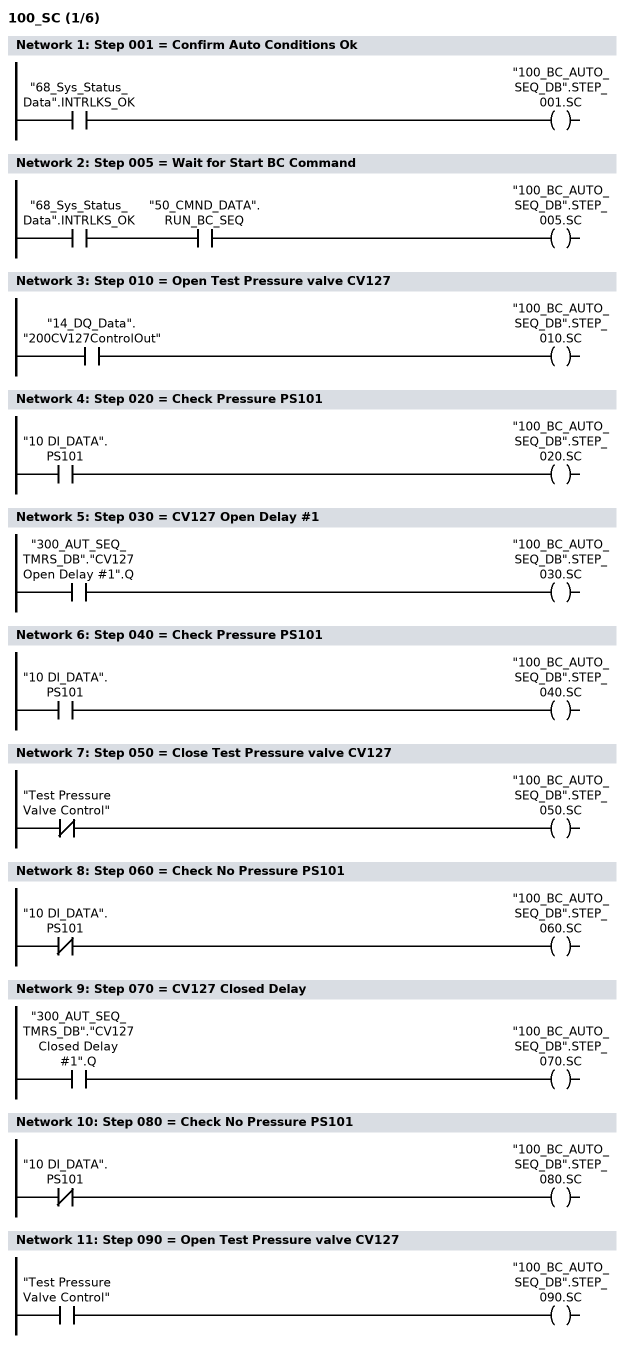
   RUNG wire#powerrail
      Contact( "68_Sys_Status_Data".INTRLKS_OK )
      Coil( "100_BC_AUTO_SEQ_DB".STEP_001.SC )
   END_RUNG
   // the same network as SCL:
   "100_BC_AUTO_SEQ_DB".STEP_001.SC := "68_Sys_Status_Data".INTRLKS_OK;
END_REGION

REGION Network 2: Step 005 = Wait for Start BC Command
   RUNG wire#powerrail
      Contact( "68_Sys_Status_Data".INTRLKS_OK )
      Contact( "50_CMND_DATA".RUN_BC_SEQ )
      Coil( "100_BC_AUTO_SEQ_DB".STEP_005.SC )
   END_RUNG
   // the same network as SCL:
   "100_BC_AUTO_SEQ_DB".STEP_005.SC := "68_Sys_Status_Data".INTRLKS_OK AND "50_CMND_DATA".RUN_BC_SEQ;
END_REGION

REGION Network 3: Step 010 = Open Test Pressure valve CV127
   RUNG wire#powerrail
      Contact( "14_DQ_Data"."200CV127ControlOut" )
      Coil( "100_BC_AUTO_SEQ_DB".STEP_010.SC )
   END_RUNG
   // the same network as SCL:
   "100_BC_AUTO_SEQ_DB".STEP_010.SC := "14_DQ_Data"."200CV127ControlOut";
END_REGION

REGION Network 4: Step 020 = Check Pressure PS101
   RUNG wire#powerrail
      Contact( "10 DI_DATA".PS101 )
      Coil( "100_BC_AUTO_SEQ_DB".STEP_020.SC )
   END_RUNG
   // the same network as SCL:
   "100_BC_AUTO_SEQ_DB".STEP_020.SC := "10 DI_DATA".PS101;
END_REGION

REGION Network 5: Step 030 = CV127 Open Delay #1
   RUNG wire#powerrail
      Contact( "300_AUT_SEQ_TMRS_DB"."CV127 Open Delay #1".Q )
      Coil( "100_BC_AUTO_SEQ_DB".STEP_030.SC )
   END_RUNG
   // the same network as SCL:
   "100_BC_AUTO_SEQ_DB".STEP_030.SC := "300_AUT_SEQ_TMRS_DB"."CV127 Open Delay #1".Q;
END_REGION

REGION Network 6: Step 040 = Check Pressure PS101
   RUNG wire#powerrail
      Contact( "10 DI_DATA".PS101 )
      Coil( "100_BC_AUTO_SEQ_DB".STEP_040.SC )
   END_RUNG
   // the same network as SCL:
   "100_BC_AUTO_SEQ_DB".STEP_040.SC := "10 DI_DATA".PS101;
END_REGION

REGION Network 7: Step 050 = Close Test Pressure valve CV127
   RUNG wire#powerrail
      I_Contact( "Test Pressure Valve Control" )
      Coil( "100_BC_AUTO_SEQ_DB".STEP_050.SC )
   END_RUNG
   // the same network as SCL:
   "100_BC_AUTO_SEQ_DB".STEP_050.SC := NOT "Test Pressure Valve Control";
END_REGION

REGION Network 8: Step 060 = Check No Pressure PS101
   RUNG wire#powerrail
      I_Contact( "10 DI_DATA".PS101 )
      Coil( "100_BC_AUTO_SEQ_DB".STEP_060.SC )
   END_RUNG
   // the same network as SCL:
   "100_BC_AUTO_SEQ_DB".STEP_060.SC := NOT "10 DI_DATA".PS101;
END_REGION

REGION Network 9: Step 070 = CV127 Closed Delay
   RUNG wire#powerrail
      Contact( "300_AUT_SEQ_TMRS_DB"."CV127 Closed Delay #1".Q )
      Coil( "100_BC_AUTO_SEQ_DB".STEP_070.SC )
   END_RUNG
   // the same network as SCL:
   "100_BC_AUTO_SEQ_DB".STEP_070.SC := "300_AUT_SEQ_TMRS_DB"."CV127 Closed Delay #1".Q;
END_REGION

REGION Network 10: Step 080 = Check No Pressure PS101
   RUNG wire#powerrail
      I_Contact( "10 DI_DATA".PS101 )
      Coil( "100_BC_AUTO_SEQ_DB".STEP_080.SC )
   END_RUNG
   // the same network as SCL:
   "100_BC_AUTO_SEQ_DB".STEP_080.SC := NOT "10 DI_DATA".PS101;
END_REGION

REGION Network 11: Step 090 = Open Test Pressure valve CV127
   RUNG wire#powerrail
      Contact( "Test Pressure Valve Control" )
      Coil( "100_BC_AUTO_SEQ_DB".STEP_090.SC )
   END_RUNG
   // the same network as SCL:
   "100_BC_AUTO_SEQ_DB".STEP_090.SC := "Test Pressure Valve Control";
END_REGION

REGION Network 12: Step 095 = Confirm CV403 Is Open
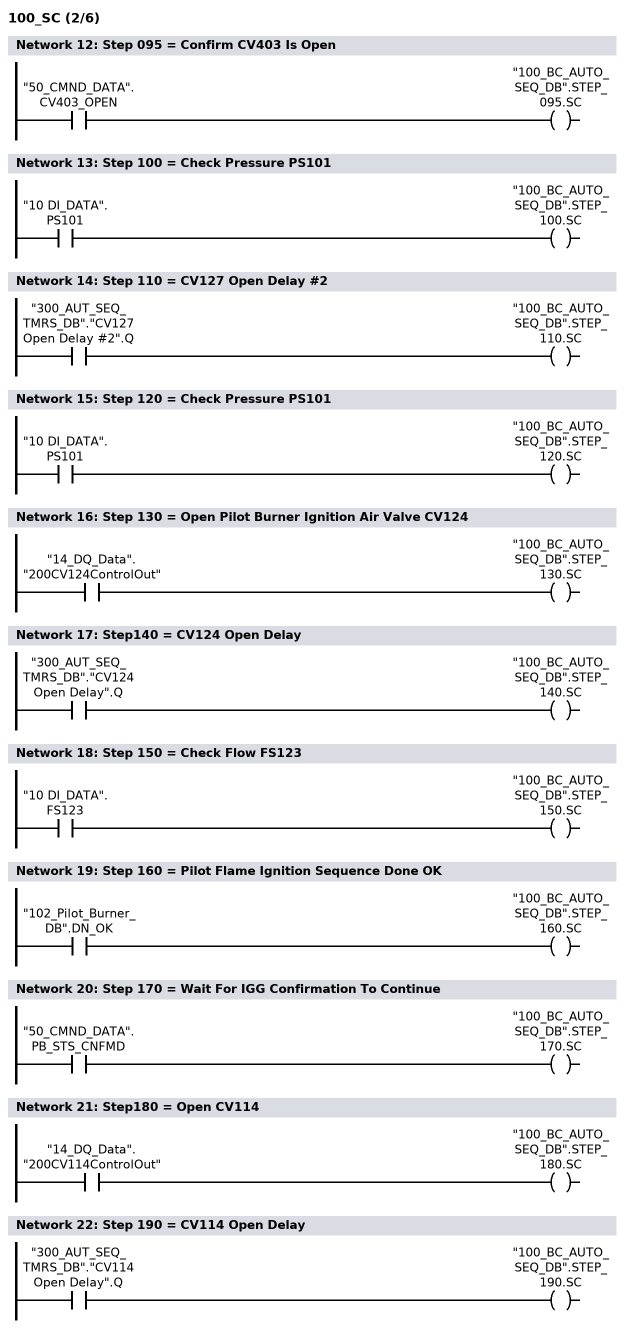
   RUNG wire#powerrail
      Contact( "50_CMND_DATA".CV403_OPEN )
      Coil( "100_BC_AUTO_SEQ_DB".STEP_095.SC )
   END_RUNG
   // the same network as SCL:
   "100_BC_AUTO_SEQ_DB".STEP_095.SC := "50_CMND_DATA".CV403_OPEN;
END_REGION

REGION Network 13: Step 100 = Check Pressure PS101
   RUNG wire#powerrail
      Contact( "10 DI_DATA".PS101 )
      Coil( "100_BC_AUTO_SEQ_DB".STEP_100.SC )
   END_RUNG
   // the same network as SCL:
   "100_BC_AUTO_SEQ_DB".STEP_100.SC := "10 DI_DATA".PS101;
END_REGION

REGION Network 14: Step 110 = CV127 Open Delay #2
   RUNG wire#powerrail
      Contact( "300_AUT_SEQ_TMRS_DB"."CV127 Open Delay #2".Q )
      Coil( "100_BC_AUTO_SEQ_DB".STEP_110.SC )
   END_RUNG
   // the same network as SCL:
   "100_BC_AUTO_SEQ_DB".STEP_110.SC := "300_AUT_SEQ_TMRS_DB"."CV127 Open Delay #2".Q;
END_REGION

REGION Network 15: Step 120 = Check Pressure PS101
   RUNG wire#powerrail
      Contact( "10 DI_DATA".PS101 )
      Coil( "100_BC_AUTO_SEQ_DB".STEP_120.SC )
   END_RUNG
   // the same network as SCL:
   "100_BC_AUTO_SEQ_DB".STEP_120.SC := "10 DI_DATA".PS101;
END_REGION

REGION Network 16: Step 130 = Open Pilot Burner Ignition Air Valve CV124
   RUNG wire#powerrail
      Contact( "14_DQ_Data"."200CV124ControlOut" )
      Coil( "100_BC_AUTO_SEQ_DB".STEP_130.SC )
   END_RUNG
   // the same network as SCL:
   "100_BC_AUTO_SEQ_DB".STEP_130.SC := "14_DQ_Data"."200CV124ControlOut";
END_REGION

REGION Network 17: Step140 = CV124 Open Delay
   RUNG wire#powerrail
      Contact( "300_AUT_SEQ_TMRS_DB"."CV124 Open Delay".Q )
      Coil( "100_BC_AUTO_SEQ_DB".STEP_140.SC )
   END_RUNG
   // the same network as SCL:
   "100_BC_AUTO_SEQ_DB".STEP_140.SC := "300_AUT_SEQ_TMRS_DB"."CV124 Open Delay".Q;
END_REGION

REGION Network 18: Step 150 = Check Flow FS123
   RUNG wire#powerrail
      Contact( "10 DI_DATA".FS123 )
      Coil( "100_BC_AUTO_SEQ_DB".STEP_150.SC )
   END_RUNG
   // the same network as SCL:
   "100_BC_AUTO_SEQ_DB".STEP_150.SC := "10 DI_DATA".FS123;
END_REGION

REGION Network 19: Step 160 = Pilot Flame Ignition Sequence Done OK
   RUNG wire#powerrail
      Contact( "102_Pilot_Burner_DB".DN_OK )
      Coil( "100_BC_AUTO_SEQ_DB".STEP_160.SC )
   END_RUNG
   // the same network as SCL:
   "100_BC_AUTO_SEQ_DB".STEP_160.SC := "102_Pilot_Burner_DB".DN_OK;
END_REGION

REGION Network 20: Step 170 = Wait For IGG Confirmation To Continue
   RUNG wire#powerrail
      Contact( "50_CMND_DATA".PB_STS_CNFMD )
      Coil( "100_BC_AUTO_SEQ_DB".STEP_170.SC )
   END_RUNG
   // the same network as SCL:
   "100_BC_AUTO_SEQ_DB".STEP_170.SC := "50_CMND_DATA".PB_STS_CNFMD;
END_REGION

REGION Network 21: Step180 = Open CV114
   RUNG wire#powerrail
      Contact( "14_DQ_Data"."200CV114ControlOut" )
      Coil( "100_BC_AUTO_SEQ_DB".STEP_180.SC )
   END_RUNG
   // the same network as SCL:
   "100_BC_AUTO_SEQ_DB".STEP_180.SC := "14_DQ_Data"."200CV114ControlOut";
END_REGION

REGION Network 22: Step 190 = CV114 Open Delay
   RUNG wire#powerrail
      Contact( "300_AUT_SEQ_TMRS_DB"."CV114 Open Delay".Q )
      Coil( "100_BC_AUTO_SEQ_DB".STEP_190.SC )
   END_RUNG
   // the same network as SCL:
   "100_BC_AUTO_SEQ_DB".STEP_190.SC := "300_AUT_SEQ_TMRS_DB"."CV114 Open Delay".Q;
END_REGION

REGION Network 23: Step 200 = Main Burner Ignition Sequence
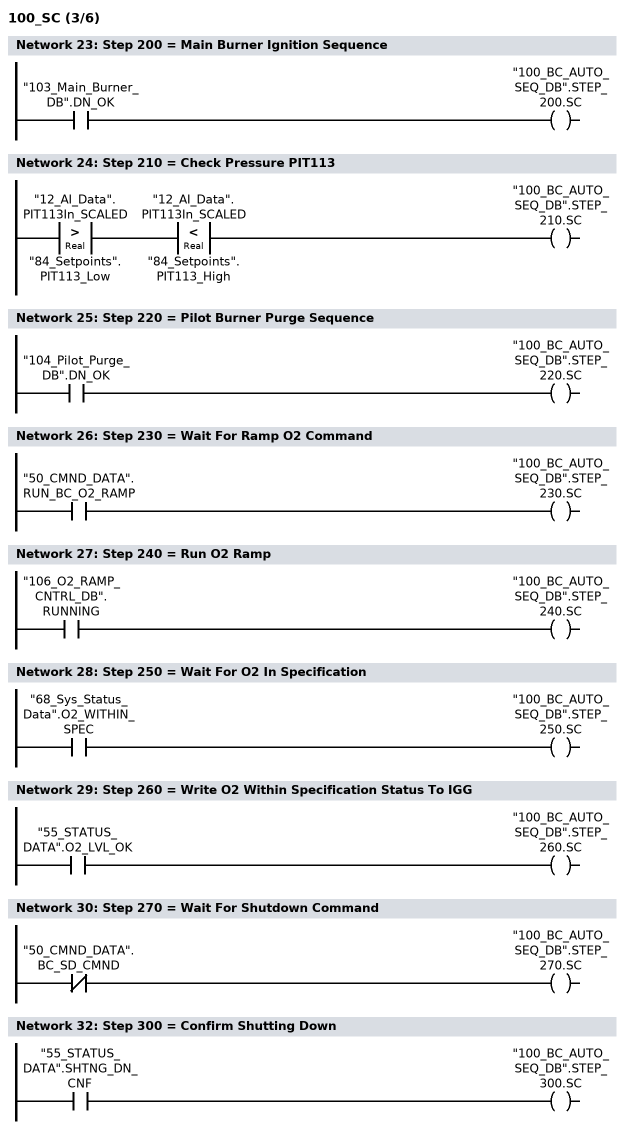
   RUNG wire#powerrail
      Contact( "103_Main_Burner_DB".DN_OK )
      Coil( "100_BC_AUTO_SEQ_DB".STEP_200.SC )
   END_RUNG
   // the same network as SCL:
   "100_BC_AUTO_SEQ_DB".STEP_200.SC := "103_Main_Burner_DB".DN_OK;
END_REGION

REGION Network 24: Step 210 = Check Pressure PIT113
   RUNG wire#powerrail
      { S7_Templates := "SrcType := Real" } GT_Contact(in1 := "12_AI_Data".PIT113In_SCALED, in2 := "84_Setpoints".PIT113_Low)
      { S7_Templates := "SrcType := Real" } LT_Contact(in1 := "12_AI_Data".PIT113In_SCALED, in2 := "84_Setpoints".PIT113_High)
      Coil( "100_BC_AUTO_SEQ_DB".STEP_210.SC )
   END_RUNG
   // the same network as SCL:
   "100_BC_AUTO_SEQ_DB".STEP_210.SC := ("12_AI_Data".PIT113In_SCALED > "84_Setpoints".PIT113_Low) AND ("12_AI_Data".PIT113In_SCALED < "84_Setpoints".PIT113_High);
END_REGION

REGION Network 25: Step 220 = Pilot Burner Purge Sequence
   RUNG wire#powerrail
      Contact( "104_Pilot_Purge_DB".DN_OK )
      Coil( "100_BC_AUTO_SEQ_DB".STEP_220.SC )
   END_RUNG
   // the same network as SCL:
   "100_BC_AUTO_SEQ_DB".STEP_220.SC := "104_Pilot_Purge_DB".DN_OK;
END_REGION

REGION Network 26: Step 230 = Wait For Ramp O2 Command
   RUNG wire#powerrail
      Contact( "50_CMND_DATA".RUN_BC_O2_RAMP )
      Coil( "100_BC_AUTO_SEQ_DB".STEP_230.SC )
   END_RUNG
   // the same network as SCL:
   "100_BC_AUTO_SEQ_DB".STEP_230.SC := "50_CMND_DATA".RUN_BC_O2_RAMP;
END_REGION

REGION Network 27: Step 240 = Run O2 Ramp
   RUNG wire#powerrail
      Contact( "106_O2_RAMP_CNTRL_DB".RUNNING )
      Coil( "100_BC_AUTO_SEQ_DB".STEP_240.SC )
   END_RUNG
   // the same network as SCL:
   "100_BC_AUTO_SEQ_DB".STEP_240.SC := "106_O2_RAMP_CNTRL_DB".RUNNING;
END_REGION

REGION Network 28: Step 250 = Wait For O2 In Specification
   RUNG wire#powerrail
      Contact( "68_Sys_Status_Data".O2_WITHIN_SPEC )
      Coil( "100_BC_AUTO_SEQ_DB".STEP_250.SC )
   END_RUNG
   // the same network as SCL:
   "100_BC_AUTO_SEQ_DB".STEP_250.SC := "68_Sys_Status_Data".O2_WITHIN_SPEC;
END_REGION

REGION Network 29: Step 260 = Write O2 Within Specification Status To IGG
   RUNG wire#powerrail
      Contact( "55_STATUS_DATA".O2_LVL_OK )
      Coil( "100_BC_AUTO_SEQ_DB".STEP_260.SC )
   END_RUNG
   // the same network as SCL:
   "100_BC_AUTO_SEQ_DB".STEP_260.SC := "55_STATUS_DATA".O2_LVL_OK;
END_REGION

REGION Network 30: Step 270 = Wait For Shutdown Command
   RUNG wire#powerrail
      I_Contact( "50_CMND_DATA".BC_SD_CMND )
      Coil( "100_BC_AUTO_SEQ_DB".STEP_270.SC )
   END_RUNG
   // the same network as SCL:
   "100_BC_AUTO_SEQ_DB".STEP_270.SC := NOT "50_CMND_DATA".BC_SD_CMND;
END_REGION

REGION Network 32: Step 300 = Confirm Shutting Down
   RUNG wire#powerrail
      Contact( "55_STATUS_DATA".SHTNG_DN_CNF )
      Coil( "100_BC_AUTO_SEQ_DB".STEP_300.SC )
   END_RUNG
   // the same network as SCL:
   "100_BC_AUTO_SEQ_DB".STEP_300.SC := "55_STATUS_DATA".SHTNG_DN_CNF;
END_REGION

REGION Network 33: Step 310 = CV203 To High O2 Standard Burn Setting
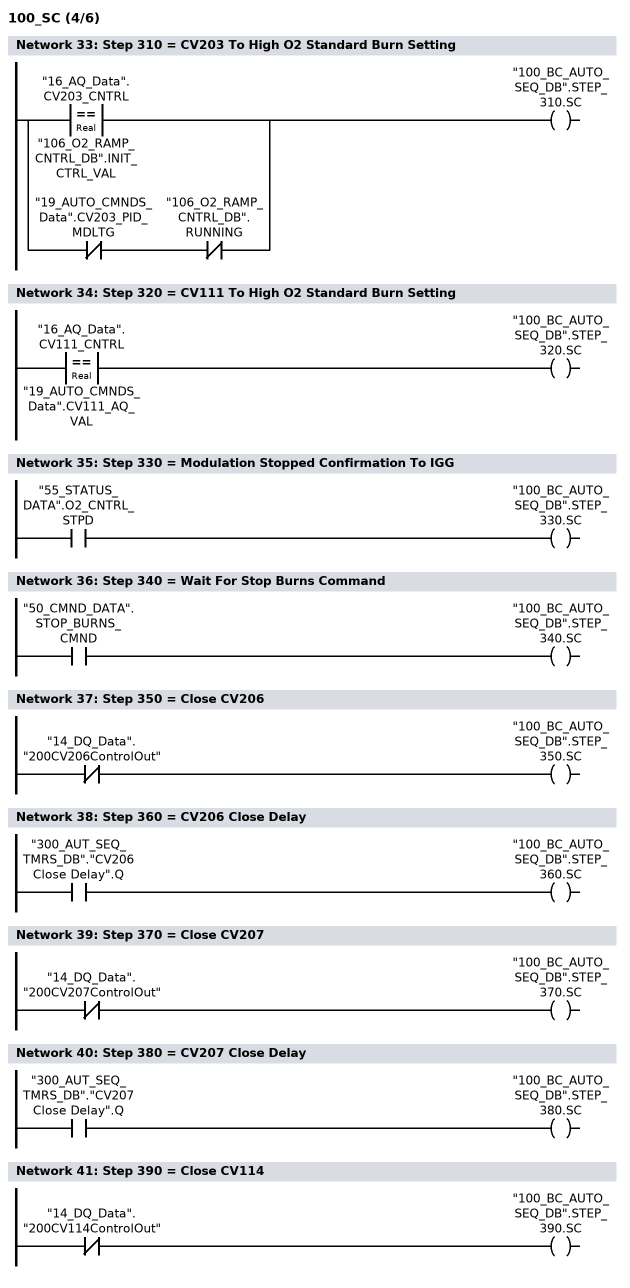
   RUNG wire#powerrail
      { S7_Templates := "SrcType := Real" } EQ_Contact(in1 := "16_AQ_Data".CV203_CNTRL, in2 := "106_O2_RAMP_CNTRL_DB".INIT_CTRL_VAL)
      wire#w1
      Coil( "100_BC_AUTO_SEQ_DB".STEP_310.SC )
   END_RUNG
   RUNG wire#powerrail
      I_Contact( "19_AUTO_CMNDS_Data".CV203_PID_MDLTG )
      I_Contact( "106_O2_RAMP_CNTRL_DB".RUNNING )
   END_RUNG wire#w1
   // the same network as SCL:
   "100_BC_AUTO_SEQ_DB".STEP_310.SC := ("16_AQ_Data".CV203_CNTRL = "106_O2_RAMP_CNTRL_DB".INIT_CTRL_VAL) OR (NOT "19_AUTO_CMNDS_Data".CV203_PID_MDLTG AND NOT "106_O2_RAMP_CNTRL_DB".RUNNING);
END_REGION

REGION Network 34: Step 320 = CV111 To High O2 Standard Burn Setting
   RUNG wire#powerrail
      { S7_Templates := "SrcType := Real" } EQ_Contact(in1 := "16_AQ_Data".CV111_CNTRL, in2 := "19_AUTO_CMNDS_Data".CV111_AQ_VAL)
      Coil( "100_BC_AUTO_SEQ_DB".STEP_320.SC )
   END_RUNG
   // the same network as SCL:
   "100_BC_AUTO_SEQ_DB".STEP_320.SC := "16_AQ_Data".CV111_CNTRL = "19_AUTO_CMNDS_Data".CV111_AQ_VAL;
END_REGION

REGION Network 35: Step 330 = Modulation Stopped Confirmation To IGG
   RUNG wire#powerrail
      Contact( "55_STATUS_DATA".O2_CNTRL_STPD )
      Coil( "100_BC_AUTO_SEQ_DB".STEP_330.SC )
   END_RUNG
   // the same network as SCL:
   "100_BC_AUTO_SEQ_DB".STEP_330.SC := "55_STATUS_DATA".O2_CNTRL_STPD;
END_REGION

REGION Network 36: Step 340 = Wait For Stop Burns Command
   RUNG wire#powerrail
      Contact( "50_CMND_DATA".STOP_BURNS_CMND )
      Coil( "100_BC_AUTO_SEQ_DB".STEP_340.SC )
   END_RUNG
   // the same network as SCL:
   "100_BC_AUTO_SEQ_DB".STEP_340.SC := "50_CMND_DATA".STOP_BURNS_CMND;
END_REGION

REGION Network 37: Step 350 = Close CV206
   RUNG wire#powerrail
      I_Contact( "14_DQ_Data"."200CV206ControlOut" )
      Coil( "100_BC_AUTO_SEQ_DB".STEP_350.SC )
   END_RUNG
   // the same network as SCL:
   "100_BC_AUTO_SEQ_DB".STEP_350.SC := NOT "14_DQ_Data"."200CV206ControlOut";
END_REGION

REGION Network 38: Step 360 = CV206 Close Delay
   RUNG wire#powerrail
      Contact( "300_AUT_SEQ_TMRS_DB"."CV206 Close Delay".Q )
      Coil( "100_BC_AUTO_SEQ_DB".STEP_360.SC )
   END_RUNG
   // the same network as SCL:
   "100_BC_AUTO_SEQ_DB".STEP_360.SC := "300_AUT_SEQ_TMRS_DB"."CV206 Close Delay".Q;
END_REGION

REGION Network 39: Step 370 = Close CV207
   RUNG wire#powerrail
      I_Contact( "14_DQ_Data"."200CV207ControlOut" )
      Coil( "100_BC_AUTO_SEQ_DB".STEP_370.SC )
   END_RUNG
   // the same network as SCL:
   "100_BC_AUTO_SEQ_DB".STEP_370.SC := NOT "14_DQ_Data"."200CV207ControlOut";
END_REGION

REGION Network 40: Step 380 = CV207 Close Delay
   RUNG wire#powerrail
      Contact( "300_AUT_SEQ_TMRS_DB"."CV207 Close Delay".Q )
      Coil( "100_BC_AUTO_SEQ_DB".STEP_380.SC )
   END_RUNG
   // the same network as SCL:
   "100_BC_AUTO_SEQ_DB".STEP_380.SC := "300_AUT_SEQ_TMRS_DB"."CV207 Close Delay".Q;
END_REGION

REGION Network 41: Step 390 = Close CV114
   RUNG wire#powerrail
      I_Contact( "14_DQ_Data"."200CV114ControlOut" )
      Coil( "100_BC_AUTO_SEQ_DB".STEP_390.SC )
   END_RUNG
   // the same network as SCL:
   "100_BC_AUTO_SEQ_DB".STEP_390.SC := NOT "14_DQ_Data"."200CV114ControlOut";
END_REGION

REGION Network 42: Step 400 = CV114 Close Delay
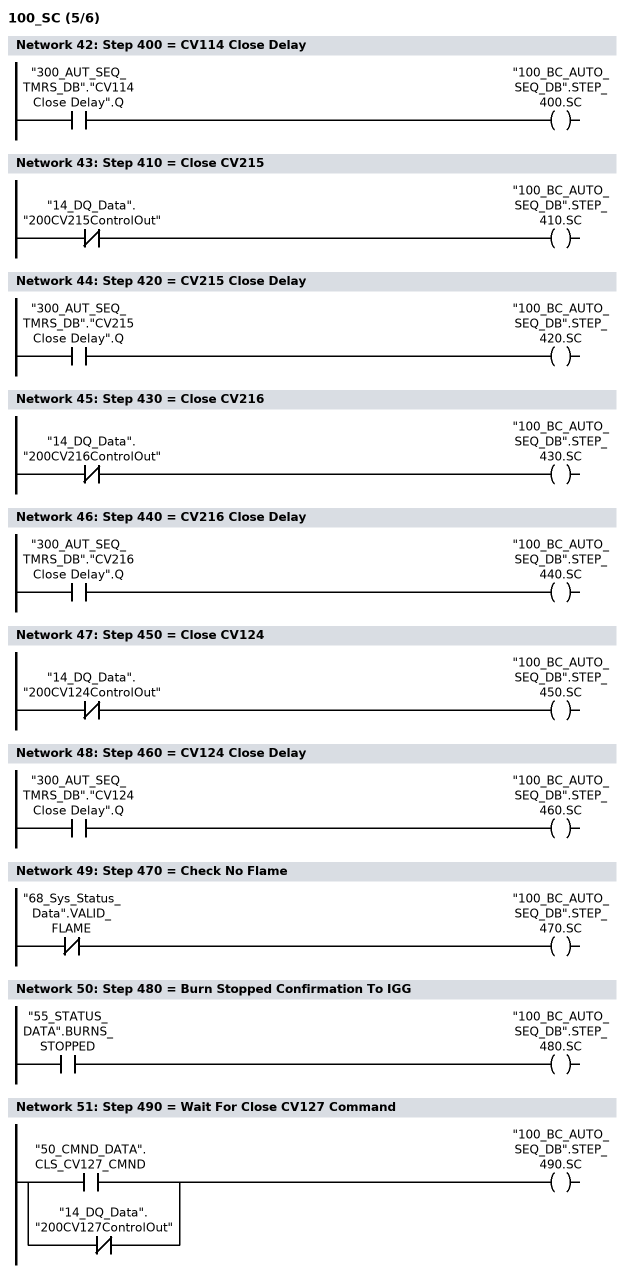
   RUNG wire#powerrail
      Contact( "300_AUT_SEQ_TMRS_DB"."CV114 Close Delay".Q )
      Coil( "100_BC_AUTO_SEQ_DB".STEP_400.SC )
   END_RUNG
   // the same network as SCL:
   "100_BC_AUTO_SEQ_DB".STEP_400.SC := "300_AUT_SEQ_TMRS_DB"."CV114 Close Delay".Q;
END_REGION

REGION Network 43: Step 410 = Close CV215
   RUNG wire#powerrail
      I_Contact( "14_DQ_Data"."200CV215ControlOut" )
      Coil( "100_BC_AUTO_SEQ_DB".STEP_410.SC )
   END_RUNG
   // the same network as SCL:
   "100_BC_AUTO_SEQ_DB".STEP_410.SC := NOT "14_DQ_Data"."200CV215ControlOut";
END_REGION

REGION Network 44: Step 420 = CV215 Close Delay
   RUNG wire#powerrail
      Contact( "300_AUT_SEQ_TMRS_DB"."CV215 Close Delay".Q )
      Coil( "100_BC_AUTO_SEQ_DB".STEP_420.SC )
   END_RUNG
   // the same network as SCL:
   "100_BC_AUTO_SEQ_DB".STEP_420.SC := "300_AUT_SEQ_TMRS_DB"."CV215 Close Delay".Q;
END_REGION

REGION Network 45: Step 430 = Close CV216
   RUNG wire#powerrail
      I_Contact( "14_DQ_Data"."200CV216ControlOut" )
      Coil( "100_BC_AUTO_SEQ_DB".STEP_430.SC )
   END_RUNG
   // the same network as SCL:
   "100_BC_AUTO_SEQ_DB".STEP_430.SC := NOT "14_DQ_Data"."200CV216ControlOut";
END_REGION

REGION Network 46: Step 440 = CV216 Close Delay
   RUNG wire#powerrail
      Contact( "300_AUT_SEQ_TMRS_DB"."CV216 Close Delay".Q )
      Coil( "100_BC_AUTO_SEQ_DB".STEP_440.SC )
   END_RUNG
   // the same network as SCL:
   "100_BC_AUTO_SEQ_DB".STEP_440.SC := "300_AUT_SEQ_TMRS_DB"."CV216 Close Delay".Q;
END_REGION

REGION Network 47: Step 450 = Close CV124
   RUNG wire#powerrail
      I_Contact( "14_DQ_Data"."200CV124ControlOut" )
      Coil( "100_BC_AUTO_SEQ_DB".STEP_450.SC )
   END_RUNG
   // the same network as SCL:
   "100_BC_AUTO_SEQ_DB".STEP_450.SC := NOT "14_DQ_Data"."200CV124ControlOut";
END_REGION

REGION Network 48: Step 460 = CV124 Close Delay
   RUNG wire#powerrail
      Contact( "300_AUT_SEQ_TMRS_DB"."CV124 Close Delay".Q )
      Coil( "100_BC_AUTO_SEQ_DB".STEP_460.SC )
   END_RUNG
   // the same network as SCL:
   "100_BC_AUTO_SEQ_DB".STEP_460.SC := "300_AUT_SEQ_TMRS_DB"."CV124 Close Delay".Q;
END_REGION

REGION Network 49: Step 470 = Check No Flame
   RUNG wire#powerrail
      I_Contact( "68_Sys_Status_Data".VALID_FLAME )
      Coil( "100_BC_AUTO_SEQ_DB".STEP_470.SC )
   END_RUNG
   // the same network as SCL:
   "100_BC_AUTO_SEQ_DB".STEP_470.SC := NOT "68_Sys_Status_Data".VALID_FLAME;
END_REGION

REGION Network 50: Step 480 = Burn Stopped Confirmation To IGG
   RUNG wire#powerrail
      Contact( "55_STATUS_DATA".BURNS_STOPPED )
      Coil( "100_BC_AUTO_SEQ_DB".STEP_480.SC )
   END_RUNG
   // the same network as SCL:
   "100_BC_AUTO_SEQ_DB".STEP_480.SC := "55_STATUS_DATA".BURNS_STOPPED;
END_REGION

REGION Network 51: Step 490 = Wait For Close CV127 Command
   RUNG wire#powerrail
      Contact( "50_CMND_DATA".CLS_CV127_CMND )
      wire#w1
      Coil( "100_BC_AUTO_SEQ_DB".STEP_490.SC )
   END_RUNG
   RUNG wire#powerrail
      I_Contact( "14_DQ_Data"."200CV127ControlOut" )
   END_RUNG wire#w1
   // the same network as SCL:
   "100_BC_AUTO_SEQ_DB".STEP_490.SC := "50_CMND_DATA".CLS_CV127_CMND OR NOT "14_DQ_Data"."200CV127ControlOut";
END_REGION

REGION Network 52: Step 500 = Close CV127
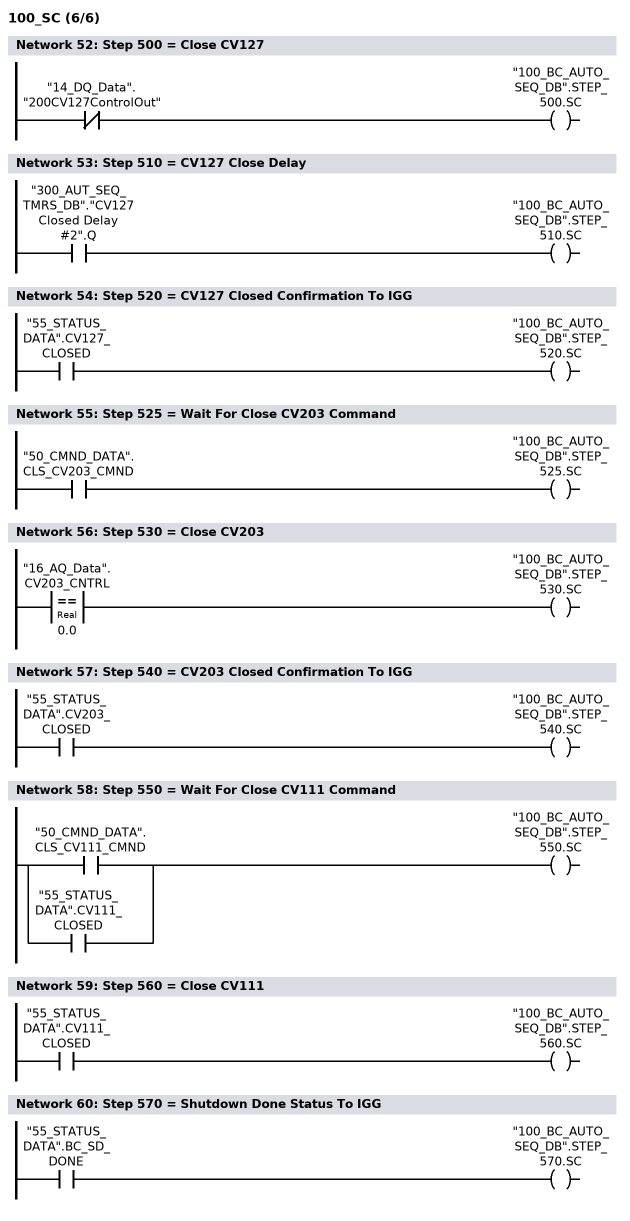
   RUNG wire#powerrail
      I_Contact( "14_DQ_Data"."200CV127ControlOut" )
      Coil( "100_BC_AUTO_SEQ_DB".STEP_500.SC )
   END_RUNG
   // the same network as SCL:
   "100_BC_AUTO_SEQ_DB".STEP_500.SC := NOT "14_DQ_Data"."200CV127ControlOut";
END_REGION

REGION Network 53: Step 510 = CV127 Close Delay
   RUNG wire#powerrail
      Contact( "300_AUT_SEQ_TMRS_DB"."CV127 Closed Delay #2".Q )
      Coil( "100_BC_AUTO_SEQ_DB".STEP_510.SC )
   END_RUNG
   // the same network as SCL:
   "100_BC_AUTO_SEQ_DB".STEP_510.SC := "300_AUT_SEQ_TMRS_DB"."CV127 Closed Delay #2".Q;
END_REGION

REGION Network 54: Step 520 = CV127 Closed Confirmation To IGG
   RUNG wire#powerrail
      Contact( "55_STATUS_DATA".CV127_CLOSED )
      Coil( "100_BC_AUTO_SEQ_DB".STEP_520.SC )
   END_RUNG
   // the same network as SCL:
   "100_BC_AUTO_SEQ_DB".STEP_520.SC := "55_STATUS_DATA".CV127_CLOSED;
END_REGION

REGION Network 55: Step 525 = Wait For Close CV203 Command
   RUNG wire#powerrail
      Contact( "50_CMND_DATA".CLS_CV203_CMND )
      Coil( "100_BC_AUTO_SEQ_DB".STEP_525.SC )
   END_RUNG
   // the same network as SCL:
   "100_BC_AUTO_SEQ_DB".STEP_525.SC := "50_CMND_DATA".CLS_CV203_CMND;
END_REGION

REGION Network 56: Step 530 = Close CV203
   RUNG wire#powerrail
      { S7_Templates := "SrcType := Real" } EQ_Contact(in1 := "16_AQ_Data".CV203_CNTRL, in2 := 0.0)
      Coil( "100_BC_AUTO_SEQ_DB".STEP_530.SC )
   END_RUNG
   // the same network as SCL:
   "100_BC_AUTO_SEQ_DB".STEP_530.SC := "16_AQ_Data".CV203_CNTRL = 0.0;
END_REGION

REGION Network 57: Step 540 = CV203 Closed Confirmation To IGG
   RUNG wire#powerrail
      Contact( "55_STATUS_DATA".CV203_CLOSED )
      Coil( "100_BC_AUTO_SEQ_DB".STEP_540.SC )
   END_RUNG
   // the same network as SCL:
   "100_BC_AUTO_SEQ_DB".STEP_540.SC := "55_STATUS_DATA".CV203_CLOSED;
END_REGION

REGION Network 58: Step 550 = Wait For Close CV111 Command
   RUNG wire#powerrail
      Contact( "50_CMND_DATA".CLS_CV111_CMND )
      wire#w1
      Coil( "100_BC_AUTO_SEQ_DB".STEP_550.SC )
   END_RUNG
   RUNG wire#powerrail
      Contact( "55_STATUS_DATA".CV111_CLOSED )
   END_RUNG wire#w1
   // the same network as SCL:
   "100_BC_AUTO_SEQ_DB".STEP_550.SC := "50_CMND_DATA".CLS_CV111_CMND OR "55_STATUS_DATA".CV111_CLOSED;
END_REGION

REGION Network 59: Step 560 = Close CV111
   RUNG wire#powerrail
      Contact( "55_STATUS_DATA".CV111_CLOSED )
      Coil( "100_BC_AUTO_SEQ_DB".STEP_560.SC )
   END_RUNG
   // the same network as SCL:
   "100_BC_AUTO_SEQ_DB".STEP_560.SC := "55_STATUS_DATA".CV111_CLOSED;
END_REGION

REGION Network 60: Step 570 = Shutdown Done Status To IGG
   RUNG wire#powerrail
      Contact( "55_STATUS_DATA".BC_SD_DONE )
      Coil( "100_BC_AUTO_SEQ_DB".STEP_570.SC )
   END_RUNG
   // the same network as SCL:
   "100_BC_AUTO_SEQ_DB".STEP_570.SC := "55_STATUS_DATA".BC_SD_DONE;
END_REGION
END_FUNCTION

// folder: 300 - 499 Counter and Timer DBs

FUNCTION "300_AUT_SUQ_TIMERS" : Void   // FC300, LAD
TITLE = Automatic Sequence Timers
{ S7_Optimized_Access := 'TRUE' }
AUTHOR : JRS
VERSION : 0.1
// For specific sequence timers not covered by step FB timers
BEGIN

REGION Network 1: Ignition Sequence Maximum Time
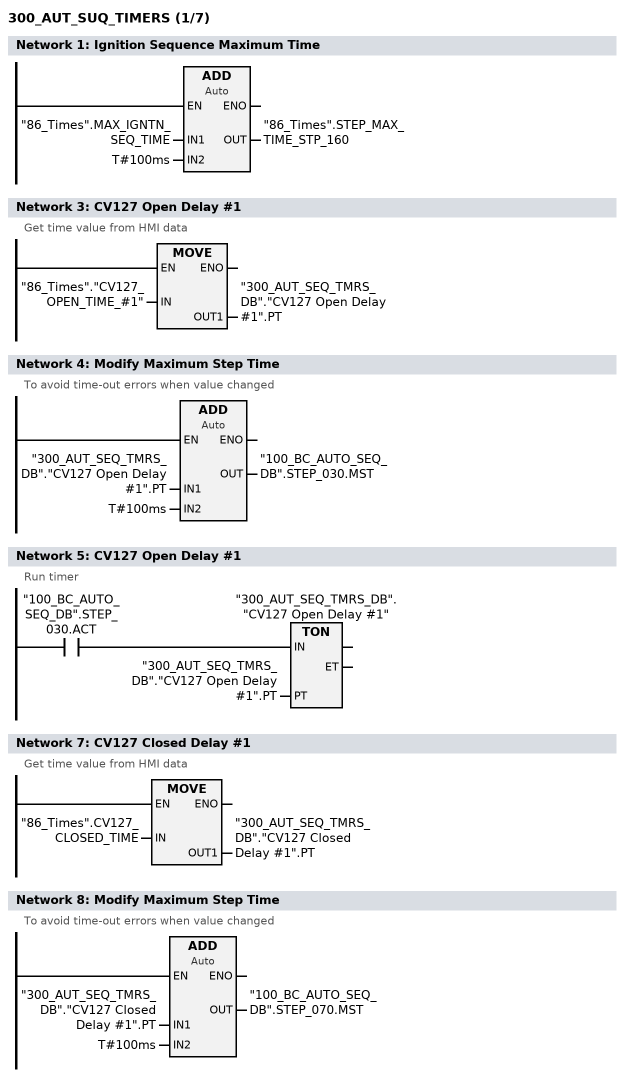
   RUNG wire#powerrail
      Add(in1 := "86_Times".MAX_IGNTN_SEQ_TIME, in2 := T#100ms, out => "86_Times".STEP_MAX_TIME_STP_160)
   END_RUNG
   // the same network as SCL:
   "86_Times".STEP_MAX_TIME_STP_160 := "86_Times".MAX_IGNTN_SEQ_TIME + T#100ms;
END_REGION

REGION Network 3: CV127 Open Delay #1
   // Get time value from HMI data
   RUNG wire#powerrail
      Move(in := "86_Times"."CV127_OPEN_TIME_#1", out1 => "300_AUT_SEQ_TMRS_DB"."CV127 Open Delay #1".PT)
   END_RUNG
   // the same network as SCL:
   "300_AUT_SEQ_TMRS_DB"."CV127 Open Delay #1".PT := "86_Times"."CV127_OPEN_TIME_#1";
END_REGION

REGION Network 4: Modify Maximum Step Time
   // To avoid time-out errors when value changed
   RUNG wire#powerrail
      Add(in1 := "300_AUT_SEQ_TMRS_DB"."CV127 Open Delay #1".PT, in2 := T#100ms, out => "100_BC_AUTO_SEQ_DB".STEP_030.MST)
   END_RUNG
   // the same network as SCL:
   "100_BC_AUTO_SEQ_DB".STEP_030.MST := "300_AUT_SEQ_TMRS_DB"."CV127 Open Delay #1".PT + T#100ms;
END_REGION

REGION Network 5: CV127 Open Delay #1
   // Run timer
   "300_AUT_SEQ_TMRS_DB"."CV127 Open Delay #1".TON(IN := "100_BC_AUTO_SEQ_DB".STEP_030.ACT,
                           PT := "300_AUT_SEQ_TMRS_DB"."CV127 Open Delay #1".PT);
END_REGION

REGION Network 7: CV127 Closed Delay #1
   // Get time value from HMI data
   RUNG wire#powerrail
      Move(in := "86_Times".CV127_CLOSED_TIME, out1 => "300_AUT_SEQ_TMRS_DB"."CV127 Closed Delay #1".PT)
   END_RUNG
   // the same network as SCL:
   "300_AUT_SEQ_TMRS_DB"."CV127 Closed Delay #1".PT := "86_Times".CV127_CLOSED_TIME;
END_REGION

REGION Network 8: Modify Maximum Step Time
   // To avoid time-out errors when value changed
   RUNG wire#powerrail
      Add(in1 := "300_AUT_SEQ_TMRS_DB"."CV127 Closed Delay #1".PT, in2 := T#100ms, out => "100_BC_AUTO_SEQ_DB".STEP_070.MST)
   END_RUNG
   // the same network as SCL:
   "100_BC_AUTO_SEQ_DB".STEP_070.MST := "300_AUT_SEQ_TMRS_DB"."CV127 Closed Delay #1".PT + T#100ms;
END_REGION

REGION Network 9: CV127 Closed Delay #1
   // Run timer
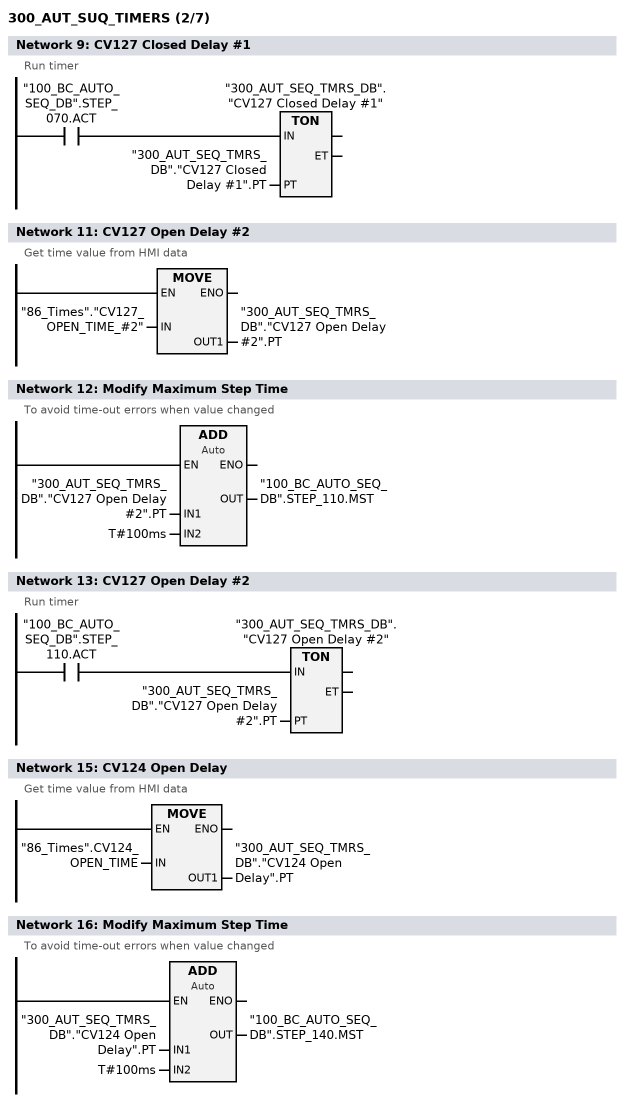
   "300_AUT_SEQ_TMRS_DB"."CV127 Closed Delay #1".TON(IN := "100_BC_AUTO_SEQ_DB".STEP_070.ACT,
                           PT := "300_AUT_SEQ_TMRS_DB"."CV127 Closed Delay #1".PT);
END_REGION

REGION Network 11: CV127 Open Delay #2
   // Get time value from HMI data
   RUNG wire#powerrail
      Move(in := "86_Times"."CV127_OPEN_TIME_#2", out1 => "300_AUT_SEQ_TMRS_DB"."CV127 Open Delay #2".PT)
   END_RUNG
   // the same network as SCL:
   "300_AUT_SEQ_TMRS_DB"."CV127 Open Delay #2".PT := "86_Times"."CV127_OPEN_TIME_#2";
END_REGION

REGION Network 12: Modify Maximum Step Time
   // To avoid time-out errors when value changed
   RUNG wire#powerrail
      Add(in1 := "300_AUT_SEQ_TMRS_DB"."CV127 Open Delay #2".PT, in2 := T#100ms, out => "100_BC_AUTO_SEQ_DB".STEP_110.MST)
   END_RUNG
   // the same network as SCL:
   "100_BC_AUTO_SEQ_DB".STEP_110.MST := "300_AUT_SEQ_TMRS_DB"."CV127 Open Delay #2".PT + T#100ms;
END_REGION

REGION Network 13: CV127 Open Delay #2
   // Run timer
   "300_AUT_SEQ_TMRS_DB"."CV127 Open Delay #2".TON(IN := "100_BC_AUTO_SEQ_DB".STEP_110.ACT,
                           PT := "300_AUT_SEQ_TMRS_DB"."CV127 Open Delay #2".PT);
END_REGION

REGION Network 15: CV124 Open Delay
   // Get time value from HMI data
   RUNG wire#powerrail
      Move(in := "86_Times".CV124_OPEN_TIME, out1 => "300_AUT_SEQ_TMRS_DB"."CV124 Open Delay".PT)
   END_RUNG
   // the same network as SCL:
   "300_AUT_SEQ_TMRS_DB"."CV124 Open Delay".PT := "86_Times".CV124_OPEN_TIME;
END_REGION

REGION Network 16: Modify Maximum Step Time
   // To avoid time-out errors when value changed
   RUNG wire#powerrail
      Add(in1 := "300_AUT_SEQ_TMRS_DB"."CV124 Open Delay".PT, in2 := T#100ms, out => "100_BC_AUTO_SEQ_DB".STEP_140.MST)
   END_RUNG
   // the same network as SCL:
   "100_BC_AUTO_SEQ_DB".STEP_140.MST := "300_AUT_SEQ_TMRS_DB"."CV124 Open Delay".PT + T#100ms;
END_REGION

REGION Network 17: CV124 Open Delay
   // Run timer
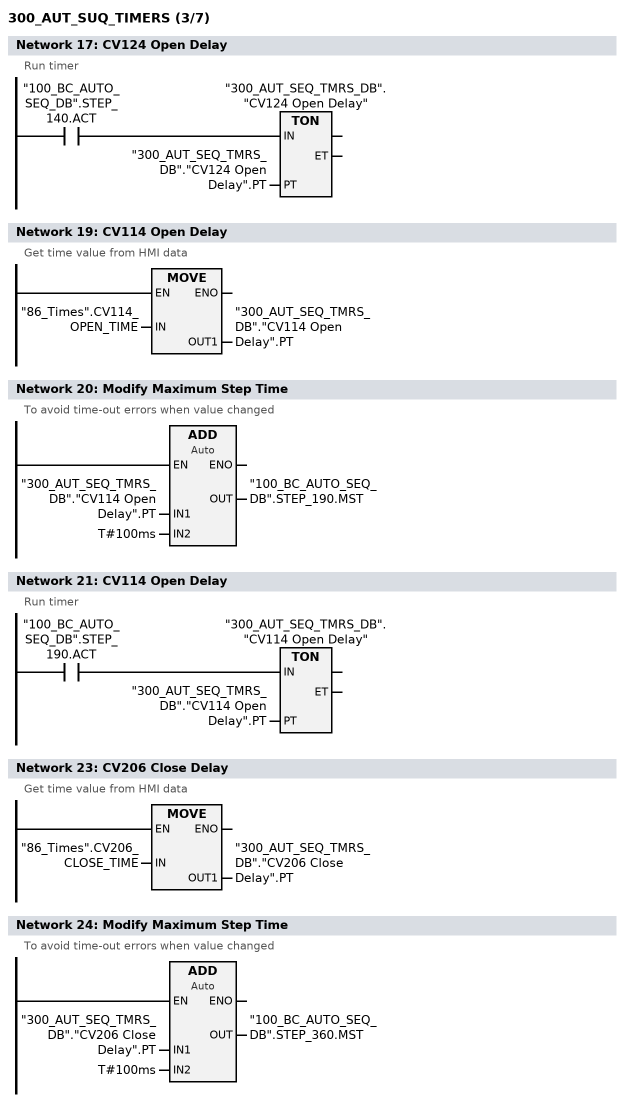
   "300_AUT_SEQ_TMRS_DB"."CV124 Open Delay".TON(IN := "100_BC_AUTO_SEQ_DB".STEP_140.ACT,
                           PT := "300_AUT_SEQ_TMRS_DB"."CV124 Open Delay".PT);
END_REGION

REGION Network 19: CV114 Open Delay
   // Get time value from HMI data
   RUNG wire#powerrail
      Move(in := "86_Times".CV114_OPEN_TIME, out1 => "300_AUT_SEQ_TMRS_DB"."CV114 Open Delay".PT)
   END_RUNG
   // the same network as SCL:
   "300_AUT_SEQ_TMRS_DB"."CV114 Open Delay".PT := "86_Times".CV114_OPEN_TIME;
END_REGION

REGION Network 20: Modify Maximum Step Time
   // To avoid time-out errors when value changed
   RUNG wire#powerrail
      Add(in1 := "300_AUT_SEQ_TMRS_DB"."CV114 Open Delay".PT, in2 := T#100ms, out => "100_BC_AUTO_SEQ_DB".STEP_190.MST)
   END_RUNG
   // the same network as SCL:
   "100_BC_AUTO_SEQ_DB".STEP_190.MST := "300_AUT_SEQ_TMRS_DB"."CV114 Open Delay".PT + T#100ms;
END_REGION

REGION Network 21: CV114 Open Delay
   // Run timer
   "300_AUT_SEQ_TMRS_DB"."CV114 Open Delay".TON(IN := "100_BC_AUTO_SEQ_DB".STEP_190.ACT,
                           PT := "300_AUT_SEQ_TMRS_DB"."CV114 Open Delay".PT);
END_REGION

REGION Network 23: CV206 Close Delay
   // Get time value from HMI data
   RUNG wire#powerrail
      Move(in := "86_Times".CV206_CLOSE_TIME, out1 => "300_AUT_SEQ_TMRS_DB"."CV206 Close Delay".PT)
   END_RUNG
   // the same network as SCL:
   "300_AUT_SEQ_TMRS_DB"."CV206 Close Delay".PT := "86_Times".CV206_CLOSE_TIME;
END_REGION

REGION Network 24: Modify Maximum Step Time
   // To avoid time-out errors when value changed
   RUNG wire#powerrail
      Add(in1 := "300_AUT_SEQ_TMRS_DB"."CV206 Close Delay".PT, in2 := T#100ms, out => "100_BC_AUTO_SEQ_DB".STEP_360.MST)
   END_RUNG
   // the same network as SCL:
   "100_BC_AUTO_SEQ_DB".STEP_360.MST := "300_AUT_SEQ_TMRS_DB"."CV206 Close Delay".PT + T#100ms;
END_REGION

REGION Network 25: CV206 Close Delay
   // Run timer
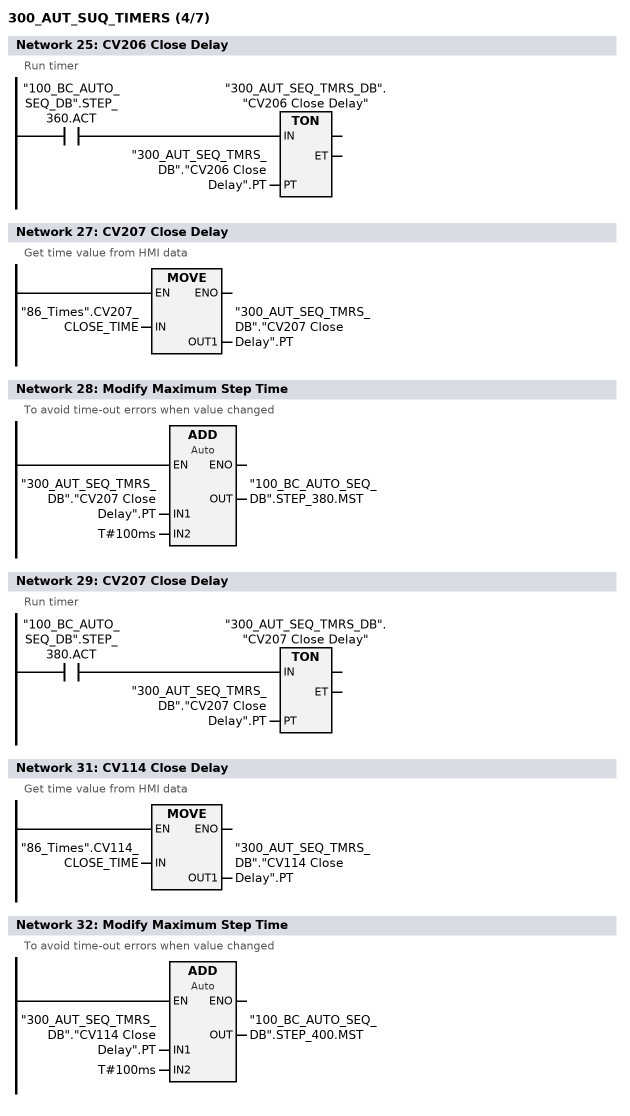
   "300_AUT_SEQ_TMRS_DB"."CV206 Close Delay".TON(IN := "100_BC_AUTO_SEQ_DB".STEP_360.ACT,
                           PT := "300_AUT_SEQ_TMRS_DB"."CV206 Close Delay".PT);
END_REGION

REGION Network 27: CV207 Close Delay
   // Get time value from HMI data
   RUNG wire#powerrail
      Move(in := "86_Times".CV207_CLOSE_TIME, out1 => "300_AUT_SEQ_TMRS_DB"."CV207 Close Delay".PT)
   END_RUNG
   // the same network as SCL:
   "300_AUT_SEQ_TMRS_DB"."CV207 Close Delay".PT := "86_Times".CV207_CLOSE_TIME;
END_REGION

REGION Network 28: Modify Maximum Step Time
   // To avoid time-out errors when value changed
   RUNG wire#powerrail
      Add(in1 := "300_AUT_SEQ_TMRS_DB"."CV207 Close Delay".PT, in2 := T#100ms, out => "100_BC_AUTO_SEQ_DB".STEP_380.MST)
   END_RUNG
   // the same network as SCL:
   "100_BC_AUTO_SEQ_DB".STEP_380.MST := "300_AUT_SEQ_TMRS_DB"."CV207 Close Delay".PT + T#100ms;
END_REGION

REGION Network 29: CV207 Close Delay
   // Run timer
   "300_AUT_SEQ_TMRS_DB"."CV207 Close Delay".TON(IN := "100_BC_AUTO_SEQ_DB".STEP_380.ACT,
                           PT := "300_AUT_SEQ_TMRS_DB"."CV207 Close Delay".PT);
END_REGION

REGION Network 31: CV114 Close Delay
   // Get time value from HMI data
   RUNG wire#powerrail
      Move(in := "86_Times".CV114_CLOSE_TIME, out1 => "300_AUT_SEQ_TMRS_DB"."CV114 Close Delay".PT)
   END_RUNG
   // the same network as SCL:
   "300_AUT_SEQ_TMRS_DB"."CV114 Close Delay".PT := "86_Times".CV114_CLOSE_TIME;
END_REGION

REGION Network 32: Modify Maximum Step Time
   // To avoid time-out errors when value changed
   RUNG wire#powerrail
      Add(in1 := "300_AUT_SEQ_TMRS_DB"."CV114 Close Delay".PT, in2 := T#100ms, out => "100_BC_AUTO_SEQ_DB".STEP_400.MST)
   END_RUNG
   // the same network as SCL:
   "100_BC_AUTO_SEQ_DB".STEP_400.MST := "300_AUT_SEQ_TMRS_DB"."CV114 Close Delay".PT + T#100ms;
END_REGION

REGION Network 33: CV114 Close Delay
   // Run timer
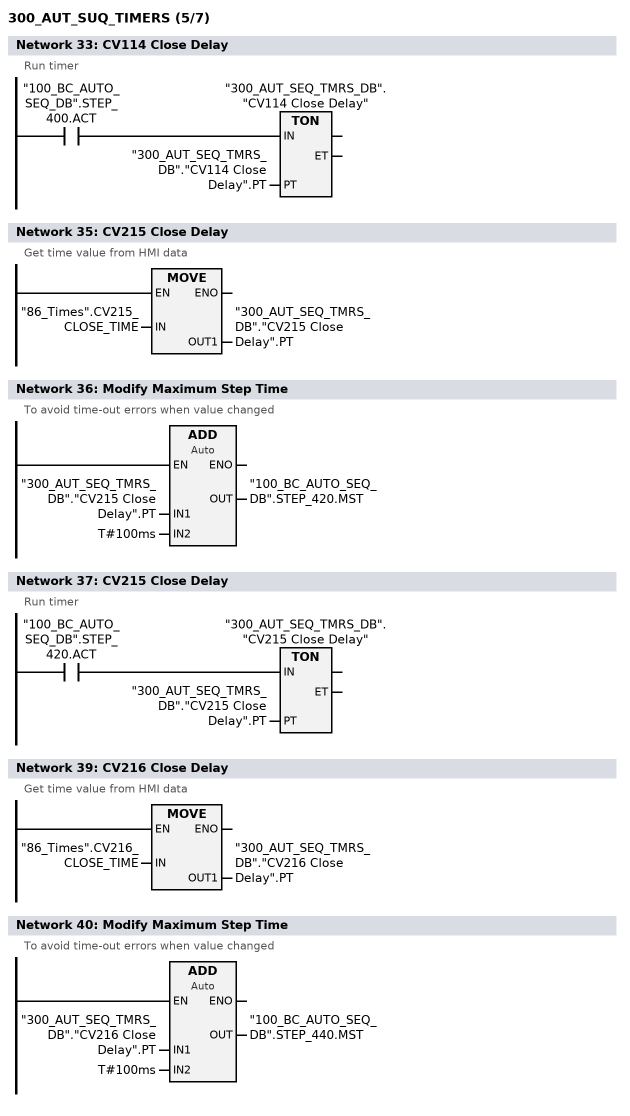
   "300_AUT_SEQ_TMRS_DB"."CV114 Close Delay".TON(IN := "100_BC_AUTO_SEQ_DB".STEP_400.ACT,
                           PT := "300_AUT_SEQ_TMRS_DB"."CV114 Close Delay".PT);
END_REGION

REGION Network 35: CV215 Close Delay
   // Get time value from HMI data
   RUNG wire#powerrail
      Move(in := "86_Times".CV215_CLOSE_TIME, out1 => "300_AUT_SEQ_TMRS_DB"."CV215 Close Delay".PT)
   END_RUNG
   // the same network as SCL:
   "300_AUT_SEQ_TMRS_DB"."CV215 Close Delay".PT := "86_Times".CV215_CLOSE_TIME;
END_REGION

REGION Network 36: Modify Maximum Step Time
   // To avoid time-out errors when value changed
   RUNG wire#powerrail
      Add(in1 := "300_AUT_SEQ_TMRS_DB"."CV215 Close Delay".PT, in2 := T#100ms, out => "100_BC_AUTO_SEQ_DB".STEP_420.MST)
   END_RUNG
   // the same network as SCL:
   "100_BC_AUTO_SEQ_DB".STEP_420.MST := "300_AUT_SEQ_TMRS_DB"."CV215 Close Delay".PT + T#100ms;
END_REGION

REGION Network 37: CV215 Close Delay
   // Run timer
   "300_AUT_SEQ_TMRS_DB"."CV215 Close Delay".TON(IN := "100_BC_AUTO_SEQ_DB".STEP_420.ACT,
                           PT := "300_AUT_SEQ_TMRS_DB"."CV215 Close Delay".PT);
END_REGION

REGION Network 39: CV216 Close Delay
   // Get time value from HMI data
   RUNG wire#powerrail
      Move(in := "86_Times".CV216_CLOSE_TIME, out1 => "300_AUT_SEQ_TMRS_DB"."CV216 Close Delay".PT)
   END_RUNG
   // the same network as SCL:
   "300_AUT_SEQ_TMRS_DB"."CV216 Close Delay".PT := "86_Times".CV216_CLOSE_TIME;
END_REGION

REGION Network 40: Modify Maximum Step Time
   // To avoid time-out errors when value changed
   RUNG wire#powerrail
      Add(in1 := "300_AUT_SEQ_TMRS_DB"."CV216 Close Delay".PT, in2 := T#100ms, out => "100_BC_AUTO_SEQ_DB".STEP_440.MST)
   END_RUNG
   // the same network as SCL:
   "100_BC_AUTO_SEQ_DB".STEP_440.MST := "300_AUT_SEQ_TMRS_DB"."CV216 Close Delay".PT + T#100ms;
END_REGION

REGION Network 41: CV216 Close Delay
   // Run timer